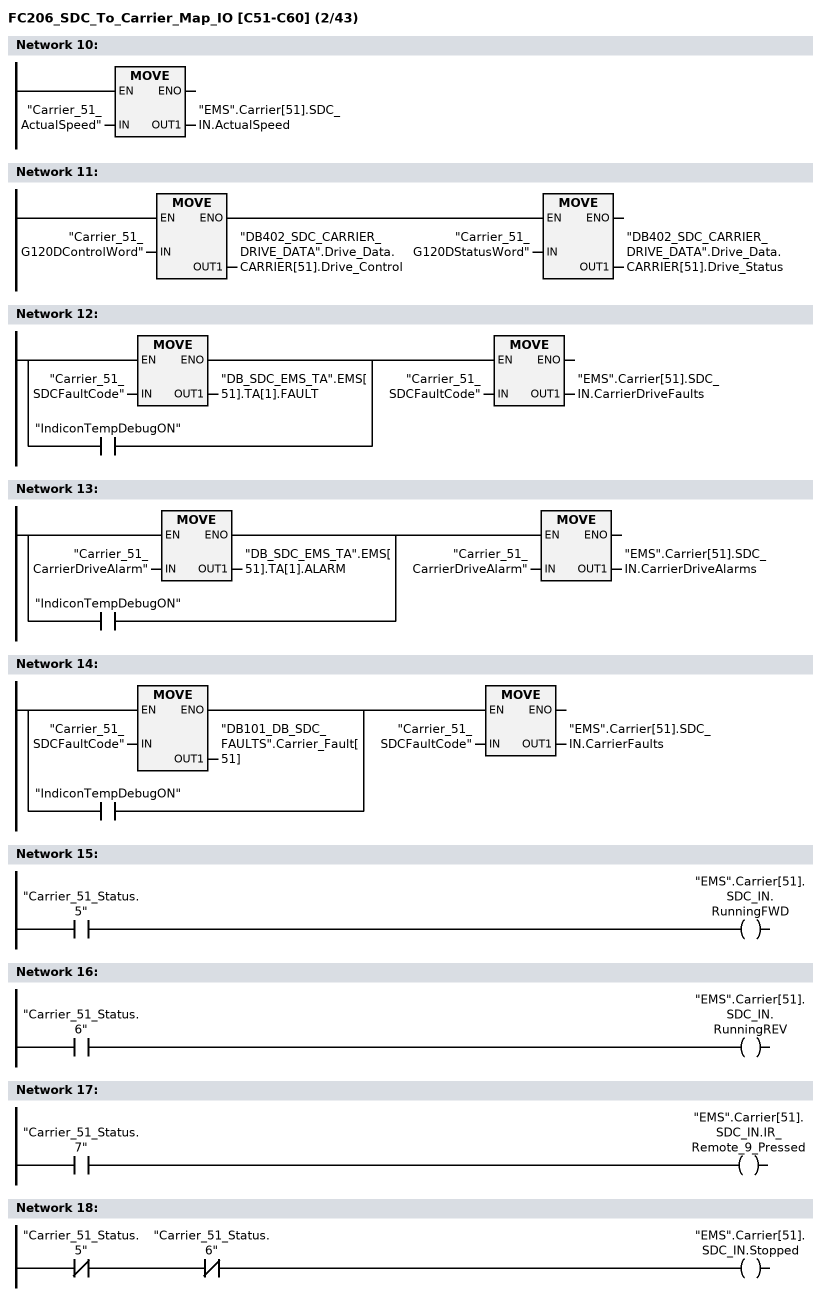
   RUNG wire#powerrail
      Move(in := "Carrier_51_ActualSpeed", out1 => "EMS".Carrier[51].SDC_IN.ActualSpeed)
   END_RUNG
   // the same network as SCL:
   "EMS".Carrier[51].SDC_IN.ActualSpeed := "Carrier_51_ActualSpeed";
END_REGION

REGION Network 11
   RUNG wire#powerrail
      Move(in := "Carrier_51_G120DControlWord", out1 => "DB402_SDC_CARRIER_DRIVE_DATA".Drive_Data.CARRIER[51].Drive_Control)
      Move(in := "Carrier_51_G120DStatusWord", out1 => "DB402_SDC_CARRIER_DRIVE_DATA".Drive_Data.CARRIER[51].Drive_Status)
   END_RUNG
   // the same network as SCL:
   "DB402_SDC_CARRIER_DRIVE_DATA".Drive_Data.CARRIER[51].Drive_Control := "Carrier_51_G120DControlWord";
   "DB402_SDC_CARRIER_DRIVE_DATA".Drive_Data.CARRIER[51].Drive_Status := "Carrier_51_G120DStatusWord";
END_REGION

REGION Network 12
   RUNG wire#powerrail
      Move(in := "Carrier_51_SDCFaultCode", out1 => "DB_SDC_EMS_TA".EMS[51].TA[1].FAULT)
      wire#w1
      Move(in := "Carrier_51_SDCFaultCode", out1 => "EMS".Carrier[51].SDC_IN.CarrierDriveFaults)
   END_RUNG
   RUNG wire#powerrail
      Contact( "IndiconTempDebugON" )
   END_RUNG wire#w1
   // the same network as SCL:
   "DB_SDC_EMS_TA".EMS[51].TA[1].FAULT := "Carrier_51_SDCFaultCode";
   IF TRUE OR "IndiconTempDebugON" THEN
       "EMS".Carrier[51].SDC_IN.CarrierDriveFaults := "Carrier_51_SDCFaultCode";
   END_IF;
END_REGION

REGION Network 13
   RUNG wire#powerrail
      Move(in := "Carrier_51_CarrierDriveAlarm", out1 => "DB_SDC_EMS_TA".EMS[51].TA[1].ALARM)
      wire#w1
      Move(in := "Carrier_51_CarrierDriveAlarm", out1 => "EMS".Carrier[51].SDC_IN.CarrierDriveAlarms)
   END_RUNG
   RUNG wire#powerrail
      Contact( "IndiconTempDebugON" )
   END_RUNG wire#w1
   // the same network as SCL:
   "DB_SDC_EMS_TA".EMS[51].TA[1].ALARM := "Carrier_51_CarrierDriveAlarm";
   IF TRUE OR "IndiconTempDebugON" THEN
       "EMS".Carrier[51].SDC_IN.CarrierDriveAlarms := "Carrier_51_CarrierDriveAlarm";
   END_IF;
END_REGION

REGION Network 14
   RUNG wire#powerrail
      Move(in := "Carrier_51_SDCFaultCode", out1 => "DB101_DB_SDC_FAULTS".Carrier_Fault[51])
      wire#w1
      Move(in := "Carrier_51_SDCFaultCode", out1 => "EMS".Carrier[51].SDC_IN.CarrierFaults)
   END_RUNG
   RUNG wire#powerrail
      Contact( "IndiconTempDebugON" )
   END_RUNG wire#w1
   // the same network as SCL:
   "DB101_DB_SDC_FAULTS".Carrier_Fault[51] := "Carrier_51_SDCFaultCode";
   IF TRUE OR "IndiconTempDebugON" THEN
       "EMS".Carrier[51].SDC_IN.CarrierFaults := "Carrier_51_SDCFaultCode";
   END_IF;
END_REGION

REGION Network 15
   RUNG wire#powerrail
      Contact( "Carrier_51_Status.5" )
      Coil( "EMS".Carrier[51].SDC_IN.RunningFWD )
   END_RUNG
   // the same network as SCL:
   "EMS".Carrier[51].SDC_IN.RunningFWD := "Carrier_51_Status.5";
END_REGION

REGION Network 16
   RUNG wire#powerrail
      Contact( "Carrier_51_Status.6" )
      Coil( "EMS".Carrier[51].SDC_IN.RunningREV )
   END_RUNG
   // the same network as SCL:
   "EMS".Carrier[51].SDC_IN.RunningREV := "Carrier_51_Status.6";
END_REGION

REGION Network 17
   RUNG wire#powerrail
      Contact( "Carrier_51_Status.7" )
      Coil( "EMS".Carrier[51].SDC_IN.IR_Remote_9_Pressed )
   END_RUNG
   // the same network as SCL:
   "EMS".Carrier[51].SDC_IN.IR_Remote_9_Pressed := "Carrier_51_Status.7";
END_REGION

REGION Network 18
   RUNG wire#powerrail
      I_Contact( "Carrier_51_Status.5" )
      I_Contact( "Carrier_51_Status.6" )
      Coil( "EMS".Carrier[51].SDC_IN.Stopped )
   END_RUNG
   // the same network as SCL:
   "EMS".Carrier[51].SDC_IN.Stopped := NOT "Carrier_51_Status.5" AND NOT "Carrier_51_Status.6";
END_REGION

REGION Network 19
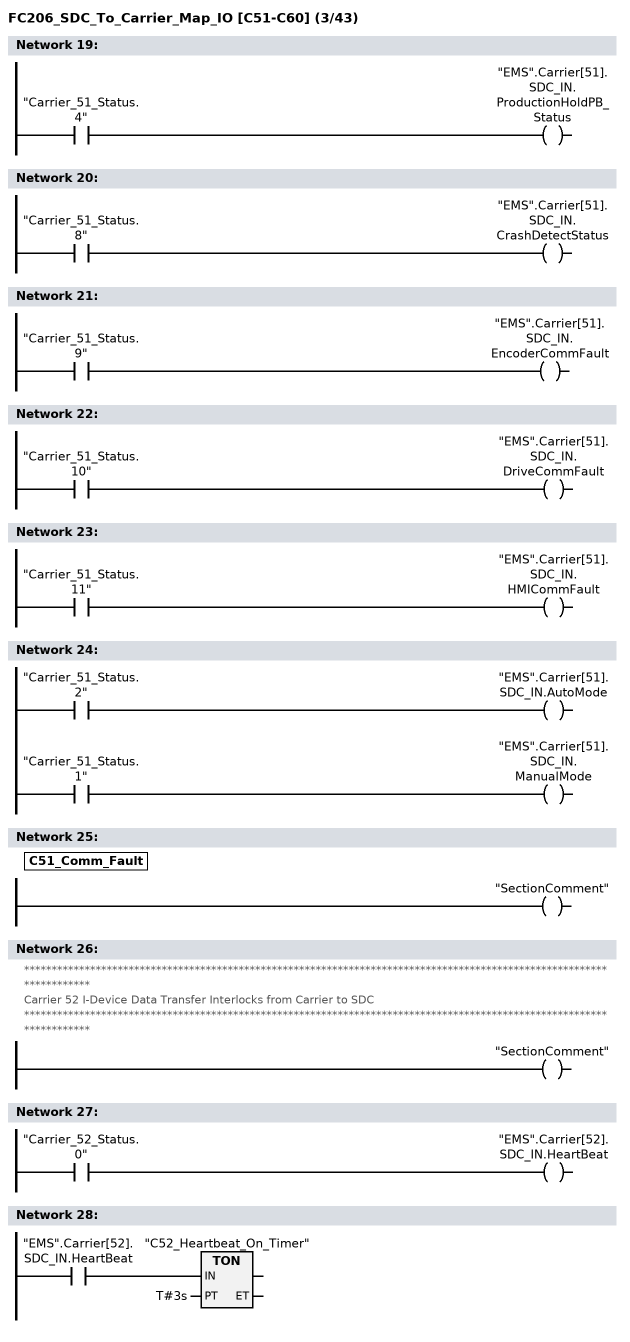
   RUNG wire#powerrail
      Contact( "Carrier_51_Status.4" )
      Coil( "EMS".Carrier[51].SDC_IN.ProductionHoldPB_Status )
   END_RUNG
   // the same network as SCL:
   "EMS".Carrier[51].SDC_IN.ProductionHoldPB_Status := "Carrier_51_Status.4";
END_REGION

REGION Network 20
   RUNG wire#powerrail
      Contact( "Carrier_51_Status.8" )
      Coil( "EMS".Carrier[51].SDC_IN.CrashDetectStatus )
   END_RUNG
   // the same network as SCL:
   "EMS".Carrier[51].SDC_IN.CrashDetectStatus := "Carrier_51_Status.8";
END_REGION

REGION Network 21
   RUNG wire#powerrail
      Contact( "Carrier_51_Status.9" )
      Coil( "EMS".Carrier[51].SDC_IN.EncoderCommFault )
   END_RUNG
   // the same network as SCL:
   "EMS".Carrier[51].SDC_IN.EncoderCommFault := "Carrier_51_Status.9";
END_REGION

REGION Network 22
   RUNG wire#powerrail
      Contact( "Carrier_51_Status.10" )
      Coil( "EMS".Carrier[51].SDC_IN.DriveCommFault )
   END_RUNG
   // the same network as SCL:
   "EMS".Carrier[51].SDC_IN.DriveCommFault := "Carrier_51_Status.10";
END_REGION

REGION Network 23
   RUNG wire#powerrail
      Contact( "Carrier_51_Status.11" )
      Coil( "EMS".Carrier[51].SDC_IN.HMICommFault )
   END_RUNG
   // the same network as SCL:
   "EMS".Carrier[51].SDC_IN.HMICommFault := "Carrier_51_Status.11";
END_REGION

REGION Network 24
   RUNG wire#powerrail
      Contact( "Carrier_51_Status.2" )
      Coil( "EMS".Carrier[51].SDC_IN.AutoMode )
   END_RUNG
   RUNG wire#powerrail
      Contact( "Carrier_51_Status.1" )
      Coil( "EMS".Carrier[51].SDC_IN.ManualMode )
   END_RUNG
   // the same network as SCL:
   "EMS".Carrier[51].SDC_IN.AutoMode := "Carrier_51_Status.2";
   "EMS".Carrier[51].SDC_IN.ManualMode := "Carrier_51_Status.1";
END_REGION

REGION Network 25
   Label( C51_Comm_Fault )
   RUNG wire#powerrail
      Coil( "SectionComment" )
   END_RUNG
   // the same network as SCL:
   C51_Comm_Fault:
   "SectionComment" := TRUE;
END_REGION

REGION Network 26
   // **********************************************************************************************************************
   // 
   // Carrier 52 I-Device Data Transfer Interlocks from Carrier to SDC
   // 
   // **********************************************************************************************************************
   RUNG wire#powerrail
      Coil( "SectionComment" )
   END_RUNG
   // the same network as SCL:
   "SectionComment" := TRUE;
END_REGION

REGION Network 27
   RUNG wire#powerrail
      Contact( "Carrier_52_Status.0" )
      Coil( "EMS".Carrier[52].SDC_IN.HeartBeat )
   END_RUNG
   // the same network as SCL:
   "EMS".Carrier[52].SDC_IN.HeartBeat := "Carrier_52_Status.0";
END_REGION

REGION Network 28
   "C52_Heartbeat_On_Timer".TON(IN := "EMS".Carrier[52].SDC_IN.HeartBeat, PT := T#3s);
END_REGION

REGION Network 29
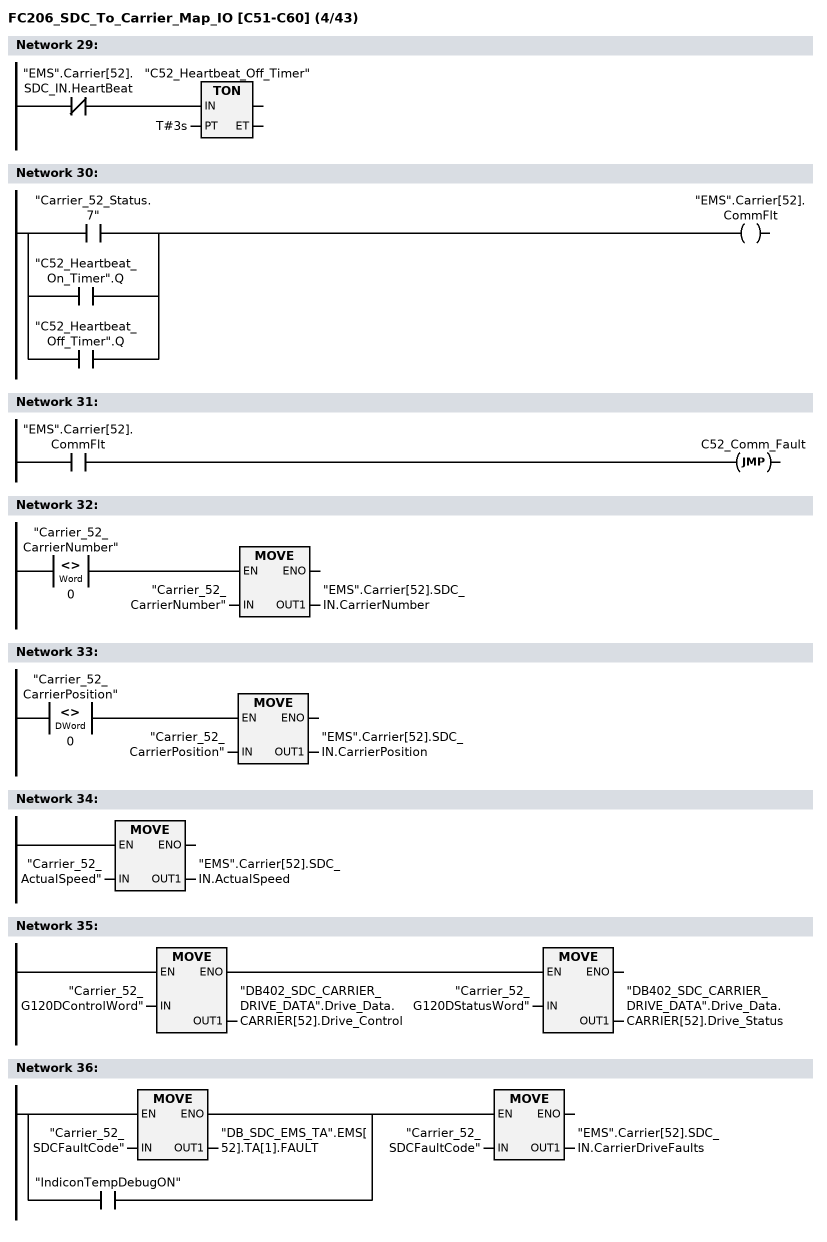
   "C52_Heartbeat_Off_Timer".TON(IN := NOT "EMS".Carrier[52].SDC_IN.HeartBeat, PT := T#3s);
END_REGION

REGION Network 30
   RUNG wire#powerrail
      Contact( "Carrier_52_Status.7" )
      wire#w1
      Coil( "EMS".Carrier[52].CommFlt )
   END_RUNG
   RUNG wire#powerrail
      Contact( "C52_Heartbeat_On_Timer".Q )
   END_RUNG wire#w1
   RUNG wire#powerrail
      Contact( "C52_Heartbeat_Off_Timer".Q )
   END_RUNG wire#w1
   // the same network as SCL:
   "EMS".Carrier[52].CommFlt := "Carrier_52_Status.7" OR "C52_Heartbeat_On_Timer".Q OR "C52_Heartbeat_Off_Timer".Q;
END_REGION

REGION Network 31
   RUNG wire#powerrail
      Contact( "EMS".Carrier[52].CommFlt )
      JumpCoil( C52_Comm_Fault )
   END_RUNG
   // the same network as SCL:
   IF "EMS".Carrier[52].CommFlt THEN GOTO C52_Comm_Fault; END_IF;
END_REGION

REGION Network 32
   RUNG wire#powerrail
      { S7_Templates := "SrcType := Word" } NE_Contact(in1 := "Carrier_52_CarrierNumber", in2 := 0)
      Move(in := "Carrier_52_CarrierNumber", out1 => "EMS".Carrier[52].SDC_IN.CarrierNumber)
   END_RUNG
   // the same network as SCL:
   IF "Carrier_52_CarrierNumber" <> 0 THEN
       "EMS".Carrier[52].SDC_IN.CarrierNumber := "Carrier_52_CarrierNumber";
   END_IF;
END_REGION

REGION Network 33
   RUNG wire#powerrail
      { S7_Templates := "SrcType := DWord" } NE_Contact(in1 := "Carrier_52_CarrierPosition", in2 := 0)
      Move(in := "Carrier_52_CarrierPosition", out1 => "EMS".Carrier[52].SDC_IN.CarrierPosition)
   END_RUNG
   // the same network as SCL:
   IF "Carrier_52_CarrierPosition" <> 0 THEN
       "EMS".Carrier[52].SDC_IN.CarrierPosition := "Carrier_52_CarrierPosition";
   END_IF;
END_REGION

REGION Network 34
   RUNG wire#powerrail
      Move(in := "Carrier_52_ActualSpeed", out1 => "EMS".Carrier[52].SDC_IN.ActualSpeed)
   END_RUNG
   // the same network as SCL:
   "EMS".Carrier[52].SDC_IN.ActualSpeed := "Carrier_52_ActualSpeed";
END_REGION

REGION Network 35
   RUNG wire#powerrail
      Move(in := "Carrier_52_G120DControlWord", out1 => "DB402_SDC_CARRIER_DRIVE_DATA".Drive_Data.CARRIER[52].Drive_Control)
      Move(in := "Carrier_52_G120DStatusWord", out1 => "DB402_SDC_CARRIER_DRIVE_DATA".Drive_Data.CARRIER[52].Drive_Status)
   END_RUNG
   // the same network as SCL:
   "DB402_SDC_CARRIER_DRIVE_DATA".Drive_Data.CARRIER[52].Drive_Control := "Carrier_52_G120DControlWord";
   "DB402_SDC_CARRIER_DRIVE_DATA".Drive_Data.CARRIER[52].Drive_Status := "Carrier_52_G120DStatusWord";
END_REGION

REGION Network 36
   RUNG wire#powerrail
      Move(in := "Carrier_52_SDCFaultCode", out1 => "DB_SDC_EMS_TA".EMS[52].TA[1].FAULT)
      wire#w1
      Move(in := "Carrier_52_SDCFaultCode", out1 => "EMS".Carrier[52].SDC_IN.CarrierDriveFaults)
   END_RUNG
   RUNG wire#powerrail
      Contact( "IndiconTempDebugON" )
   END_RUNG wire#w1
   // the same network as SCL:
   "DB_SDC_EMS_TA".EMS[52].TA[1].FAULT := "Carrier_52_SDCFaultCode";
   IF TRUE OR "IndiconTempDebugON" THEN
       "EMS".Carrier[52].SDC_IN.CarrierDriveFaults := "Carrier_52_SDCFaultCode";
   END_IF;
END_REGION

REGION Network 37
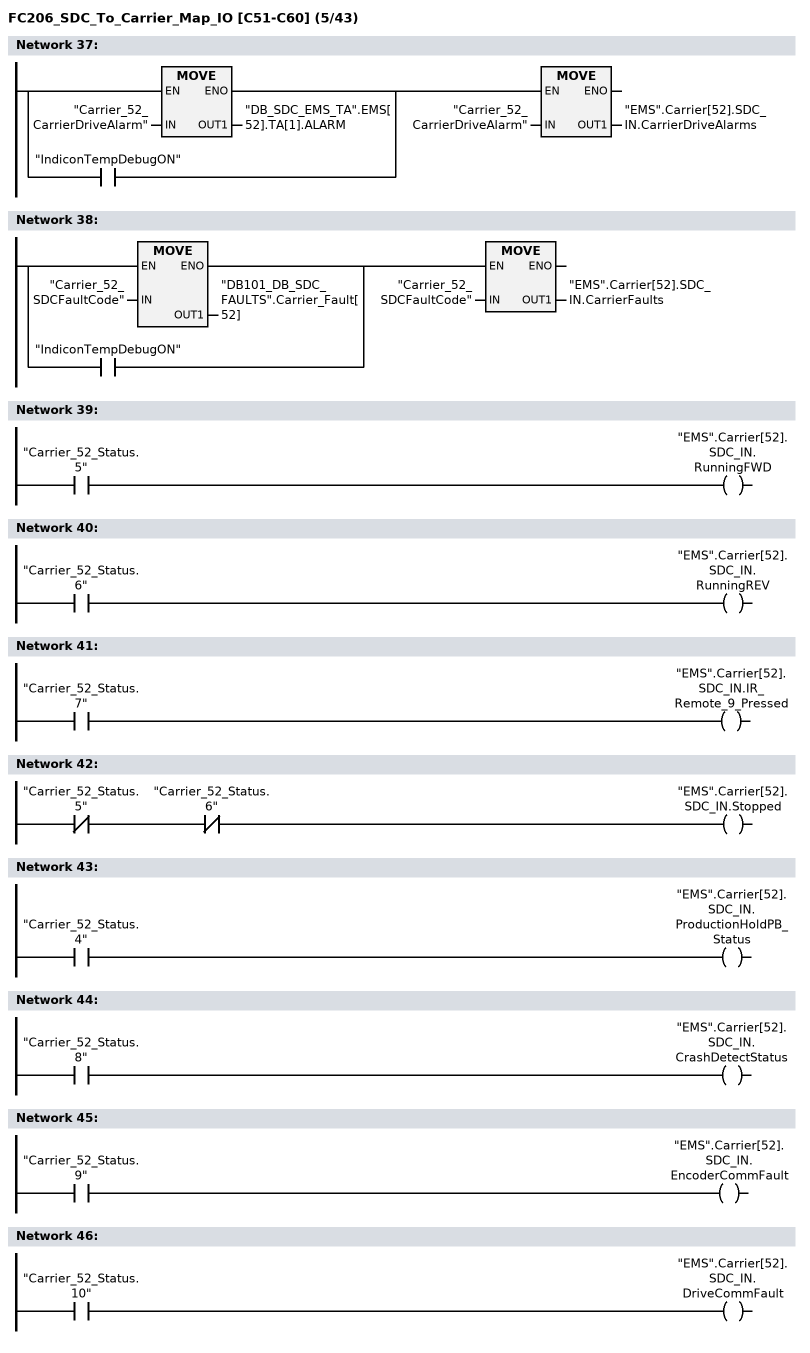
   RUNG wire#powerrail
      Move(in := "Carrier_52_CarrierDriveAlarm", out1 => "DB_SDC_EMS_TA".EMS[52].TA[1].ALARM)
      wire#w1
      Move(in := "Carrier_52_CarrierDriveAlarm", out1 => "EMS".Carrier[52].SDC_IN.CarrierDriveAlarms)
   END_RUNG
   RUNG wire#powerrail
      Contact( "IndiconTempDebugON" )
   END_RUNG wire#w1
   // the same network as SCL:
   "DB_SDC_EMS_TA".EMS[52].TA[1].ALARM := "Carrier_52_CarrierDriveAlarm";
   IF TRUE OR "IndiconTempDebugON" THEN
       "EMS".Carrier[52].SDC_IN.CarrierDriveAlarms := "Carrier_52_CarrierDriveAlarm";
   END_IF;
END_REGION

REGION Network 38
   RUNG wire#powerrail
      Move(in := "Carrier_52_SDCFaultCode", out1 => "DB101_DB_SDC_FAULTS".Carrier_Fault[52])
      wire#w1
      Move(in := "Carrier_52_SDCFaultCode", out1 => "EMS".Carrier[52].SDC_IN.CarrierFaults)
   END_RUNG
   RUNG wire#powerrail
      Contact( "IndiconTempDebugON" )
   END_RUNG wire#w1
   // the same network as SCL:
   "DB101_DB_SDC_FAULTS".Carrier_Fault[52] := "Carrier_52_SDCFaultCode";
   IF TRUE OR "IndiconTempDebugON" THEN
       "EMS".Carrier[52].SDC_IN.CarrierFaults := "Carrier_52_SDCFaultCode";
   END_IF;
END_REGION

REGION Network 39
   RUNG wire#powerrail
      Contact( "Carrier_52_Status.5" )
      Coil( "EMS".Carrier[52].SDC_IN.RunningFWD )
   END_RUNG
   // the same network as SCL:
   "EMS".Carrier[52].SDC_IN.RunningFWD := "Carrier_52_Status.5";
END_REGION

REGION Network 40
   RUNG wire#powerrail
      Contact( "Carrier_52_Status.6" )
      Coil( "EMS".Carrier[52].SDC_IN.RunningREV )
   END_RUNG
   // the same network as SCL:
   "EMS".Carrier[52].SDC_IN.RunningREV := "Carrier_52_Status.6";
END_REGION

REGION Network 41
   RUNG wire#powerrail
      Contact( "Carrier_52_Status.7" )
      Coil( "EMS".Carrier[52].SDC_IN.IR_Remote_9_Pressed )
   END_RUNG
   // the same network as SCL:
   "EMS".Carrier[52].SDC_IN.IR_Remote_9_Pressed := "Carrier_52_Status.7";
END_REGION

REGION Network 42
   RUNG wire#powerrail
      I_Contact( "Carrier_52_Status.5" )
      I_Contact( "Carrier_52_Status.6" )
      Coil( "EMS".Carrier[52].SDC_IN.Stopped )
   END_RUNG
   // the same network as SCL:
   "EMS".Carrier[52].SDC_IN.Stopped := NOT "Carrier_52_Status.5" AND NOT "Carrier_52_Status.6";
END_REGION

REGION Network 43
   RUNG wire#powerrail
      Contact( "Carrier_52_Status.4" )
      Coil( "EMS".Carrier[52].SDC_IN.ProductionHoldPB_Status )
   END_RUNG
   // the same network as SCL:
   "EMS".Carrier[52].SDC_IN.ProductionHoldPB_Status := "Carrier_52_Status.4";
END_REGION

REGION Network 44
   RUNG wire#powerrail
      Contact( "Carrier_52_Status.8" )
      Coil( "EMS".Carrier[52].SDC_IN.CrashDetectStatus )
   END_RUNG
   // the same network as SCL:
   "EMS".Carrier[52].SDC_IN.CrashDetectStatus := "Carrier_52_Status.8";
END_REGION

REGION Network 45
   RUNG wire#powerrail
      Contact( "Carrier_52_Status.9" )
      Coil( "EMS".Carrier[52].SDC_IN.EncoderCommFault )
   END_RUNG
   // the same network as SCL:
   "EMS".Carrier[52].SDC_IN.EncoderCommFault := "Carrier_52_Status.9";
END_REGION

REGION Network 46
   RUNG wire#powerrail
      Contact( "Carrier_52_Status.10" )
      Coil( "EMS".Carrier[52].SDC_IN.DriveCommFault )
   END_RUNG
   // the same network as SCL:
   "EMS".Carrier[52].SDC_IN.DriveCommFault := "Carrier_52_Status.10";
END_REGION

REGION Network 47
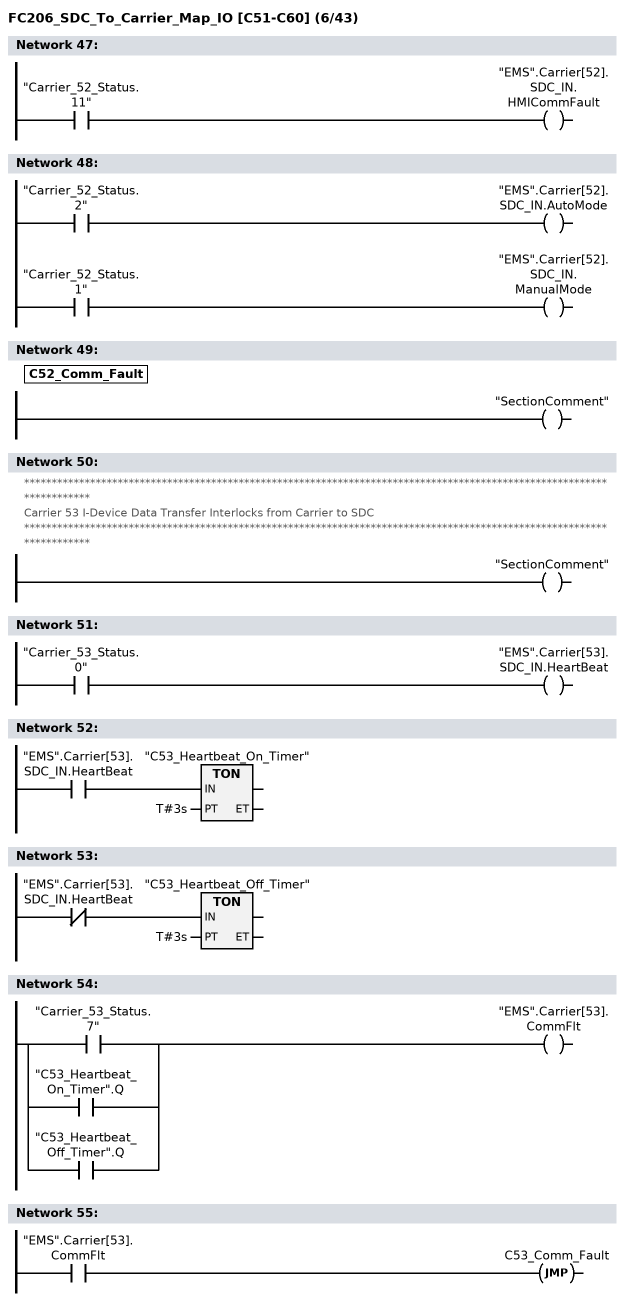
   RUNG wire#powerrail
      Contact( "Carrier_52_Status.11" )
      Coil( "EMS".Carrier[52].SDC_IN.HMICommFault )
   END_RUNG
   // the same network as SCL:
   "EMS".Carrier[52].SDC_IN.HMICommFault := "Carrier_52_Status.11";
END_REGION

REGION Network 48
   RUNG wire#powerrail
      Contact( "Carrier_52_Status.2" )
      Coil( "EMS".Carrier[52].SDC_IN.AutoMode )
   END_RUNG
   RUNG wire#powerrail
      Contact( "Carrier_52_Status.1" )
      Coil( "EMS".Carrier[52].SDC_IN.ManualMode )
   END_RUNG
   // the same network as SCL:
   "EMS".Carrier[52].SDC_IN.AutoMode := "Carrier_52_Status.2";
   "EMS".Carrier[52].SDC_IN.ManualMode := "Carrier_52_Status.1";
END_REGION

REGION Network 49
   Label( C52_Comm_Fault )
   RUNG wire#powerrail
      Coil( "SectionComment" )
   END_RUNG
   // the same network as SCL:
   C52_Comm_Fault:
   "SectionComment" := TRUE;
END_REGION

REGION Network 50
   // **********************************************************************************************************************
   // 
   // Carrier 53 I-Device Data Transfer Interlocks from Carrier to SDC
   // 
   // **********************************************************************************************************************
   RUNG wire#powerrail
      Coil( "SectionComment" )
   END_RUNG
   // the same network as SCL:
   "SectionComment" := TRUE;
END_REGION

REGION Network 51
   RUNG wire#powerrail
      Contact( "Carrier_53_Status.0" )
      Coil( "EMS".Carrier[53].SDC_IN.HeartBeat )
   END_RUNG
   // the same network as SCL:
   "EMS".Carrier[53].SDC_IN.HeartBeat := "Carrier_53_Status.0";
END_REGION

REGION Network 52
   "C53_Heartbeat_On_Timer".TON(IN := "EMS".Carrier[53].SDC_IN.HeartBeat, PT := T#3s);
END_REGION

REGION Network 53
   "C53_Heartbeat_Off_Timer".TON(IN := NOT "EMS".Carrier[53].SDC_IN.HeartBeat, PT := T#3s);
END_REGION

REGION Network 54
   RUNG wire#powerrail
      Contact( "Carrier_53_Status.7" )
      wire#w1
      Coil( "EMS".Carrier[53].CommFlt )
   END_RUNG
   RUNG wire#powerrail
      Contact( "C53_Heartbeat_On_Timer".Q )
   END_RUNG wire#w1
   RUNG wire#powerrail
      Contact( "C53_Heartbeat_Off_Timer".Q )
   END_RUNG wire#w1
   // the same network as SCL:
   "EMS".Carrier[53].CommFlt := "Carrier_53_Status.7" OR "C53_Heartbeat_On_Timer".Q OR "C53_Heartbeat_Off_Timer".Q;
END_REGION

REGION Network 55
   RUNG wire#powerrail
      Contact( "EMS".Carrier[53].CommFlt )
      JumpCoil( C53_Comm_Fault )
   END_RUNG
   // the same network as SCL:
   IF "EMS".Carrier[53].CommFlt THEN GOTO C53_Comm_Fault; END_IF;
END_REGION

REGION Network 56
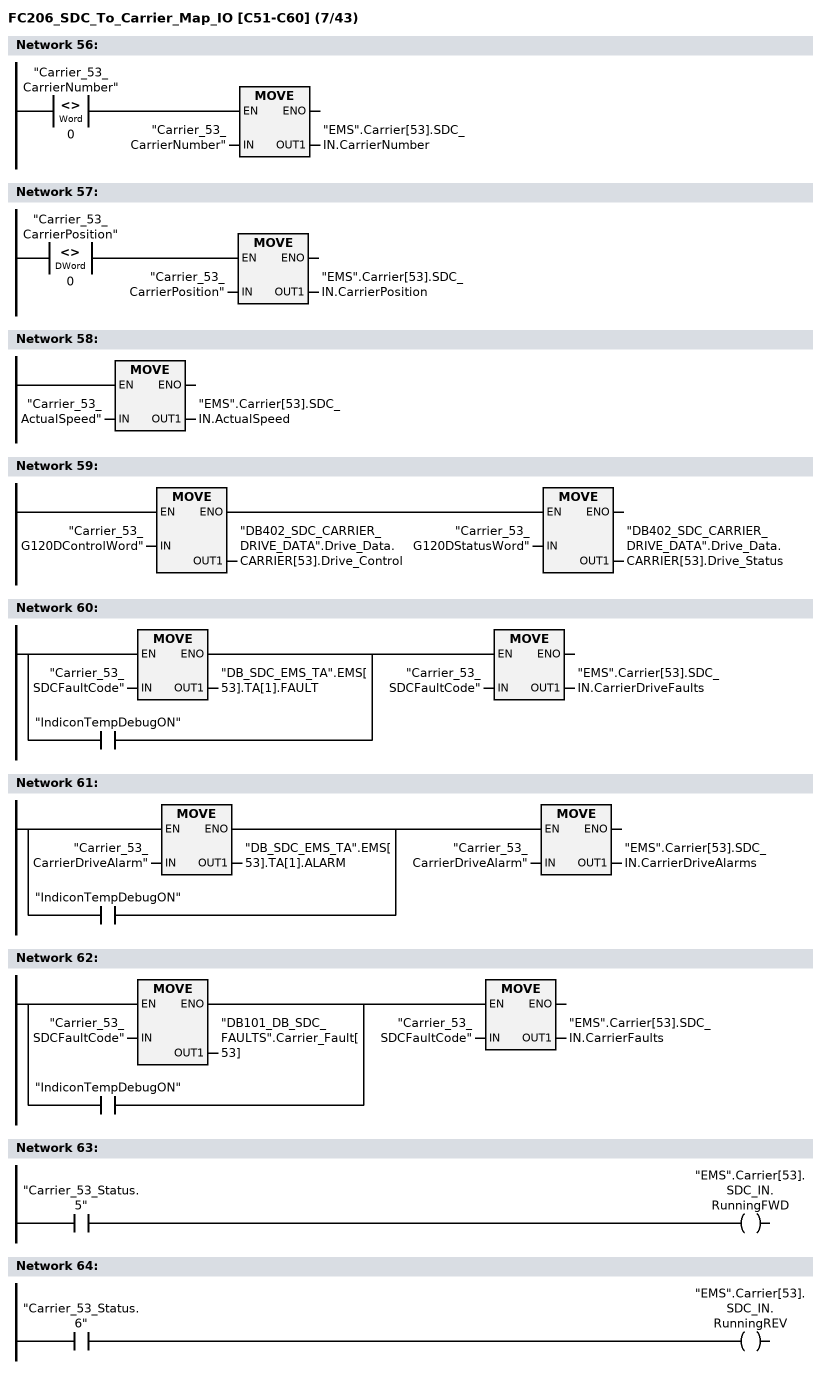
   RUNG wire#powerrail
      { S7_Templates := "SrcType := Word" } NE_Contact(in1 := "Carrier_53_CarrierNumber", in2 := 0)
      Move(in := "Carrier_53_CarrierNumber", out1 => "EMS".Carrier[53].SDC_IN.CarrierNumber)
   END_RUNG
   // the same network as SCL:
   IF "Carrier_53_CarrierNumber" <> 0 THEN
       "EMS".Carrier[53].SDC_IN.CarrierNumber := "Carrier_53_CarrierNumber";
   END_IF;
END_REGION

REGION Network 57
   RUNG wire#powerrail
      { S7_Templates := "SrcType := DWord" } NE_Contact(in1 := "Carrier_53_CarrierPosition", in2 := 0)
      Move(in := "Carrier_53_CarrierPosition", out1 => "EMS".Carrier[53].SDC_IN.CarrierPosition)
   END_RUNG
   // the same network as SCL:
   IF "Carrier_53_CarrierPosition" <> 0 THEN
       "EMS".Carrier[53].SDC_IN.CarrierPosition := "Carrier_53_CarrierPosition";
   END_IF;
END_REGION

REGION Network 58
   RUNG wire#powerrail
      Move(in := "Carrier_53_ActualSpeed", out1 => "EMS".Carrier[53].SDC_IN.ActualSpeed)
   END_RUNG
   // the same network as SCL:
   "EMS".Carrier[53].SDC_IN.ActualSpeed := "Carrier_53_ActualSpeed";
END_REGION

REGION Network 59
   RUNG wire#powerrail
      Move(in := "Carrier_53_G120DControlWord", out1 => "DB402_SDC_CARRIER_DRIVE_DATA".Drive_Data.CARRIER[53].Drive_Control)
      Move(in := "Carrier_53_G120DStatusWord", out1 => "DB402_SDC_CARRIER_DRIVE_DATA".Drive_Data.CARRIER[53].Drive_Status)
   END_RUNG
   // the same network as SCL:
   "DB402_SDC_CARRIER_DRIVE_DATA".Drive_Data.CARRIER[53].Drive_Control := "Carrier_53_G120DControlWord";
   "DB402_SDC_CARRIER_DRIVE_DATA".Drive_Data.CARRIER[53].Drive_Status := "Carrier_53_G120DStatusWord";
END_REGION

REGION Network 60
   RUNG wire#powerrail
      Move(in := "Carrier_53_SDCFaultCode", out1 => "DB_SDC_EMS_TA".EMS[53].TA[1].FAULT)
      wire#w1
      Move(in := "Carrier_53_SDCFaultCode", out1 => "EMS".Carrier[53].SDC_IN.CarrierDriveFaults)
   END_RUNG
   RUNG wire#powerrail
      Contact( "IndiconTempDebugON" )
   END_RUNG wire#w1
   // the same network as SCL:
   "DB_SDC_EMS_TA".EMS[53].TA[1].FAULT := "Carrier_53_SDCFaultCode";
   IF TRUE OR "IndiconTempDebugON" THEN
       "EMS".Carrier[53].SDC_IN.CarrierDriveFaults := "Carrier_53_SDCFaultCode";
   END_IF;
END_REGION

REGION Network 61
   RUNG wire#powerrail
      Move(in := "Carrier_53_CarrierDriveAlarm", out1 => "DB_SDC_EMS_TA".EMS[53].TA[1].ALARM)
      wire#w1
      Move(in := "Carrier_53_CarrierDriveAlarm", out1 => "EMS".Carrier[53].SDC_IN.CarrierDriveAlarms)
   END_RUNG
   RUNG wire#powerrail
      Contact( "IndiconTempDebugON" )
   END_RUNG wire#w1
   // the same network as SCL:
   "DB_SDC_EMS_TA".EMS[53].TA[1].ALARM := "Carrier_53_CarrierDriveAlarm";
   IF TRUE OR "IndiconTempDebugON" THEN
       "EMS".Carrier[53].SDC_IN.CarrierDriveAlarms := "Carrier_53_CarrierDriveAlarm";
   END_IF;
END_REGION

REGION Network 62
   RUNG wire#powerrail
      Move(in := "Carrier_53_SDCFaultCode", out1 => "DB101_DB_SDC_FAULTS".Carrier_Fault[53])
      wire#w1
      Move(in := "Carrier_53_SDCFaultCode", out1 => "EMS".Carrier[53].SDC_IN.CarrierFaults)
   END_RUNG
   RUNG wire#powerrail
      Contact( "IndiconTempDebugON" )
   END_RUNG wire#w1
   // the same network as SCL:
   "DB101_DB_SDC_FAULTS".Carrier_Fault[53] := "Carrier_53_SDCFaultCode";
   IF TRUE OR "IndiconTempDebugON" THEN
       "EMS".Carrier[53].SDC_IN.CarrierFaults := "Carrier_53_SDCFaultCode";
   END_IF;
END_REGION

REGION Network 63
   RUNG wire#powerrail
      Contact( "Carrier_53_Status.5" )
      Coil( "EMS".Carrier[53].SDC_IN.RunningFWD )
   END_RUNG
   // the same network as SCL:
   "EMS".Carrier[53].SDC_IN.RunningFWD := "Carrier_53_Status.5";
END_REGION

REGION Network 64
   RUNG wire#powerrail
      Contact( "Carrier_53_Status.6" )
      Coil( "EMS".Carrier[53].SDC_IN.RunningREV )
   END_RUNG
   // the same network as SCL:
   "EMS".Carrier[53].SDC_IN.RunningREV := "Carrier_53_Status.6";
END_REGION

REGION Network 65
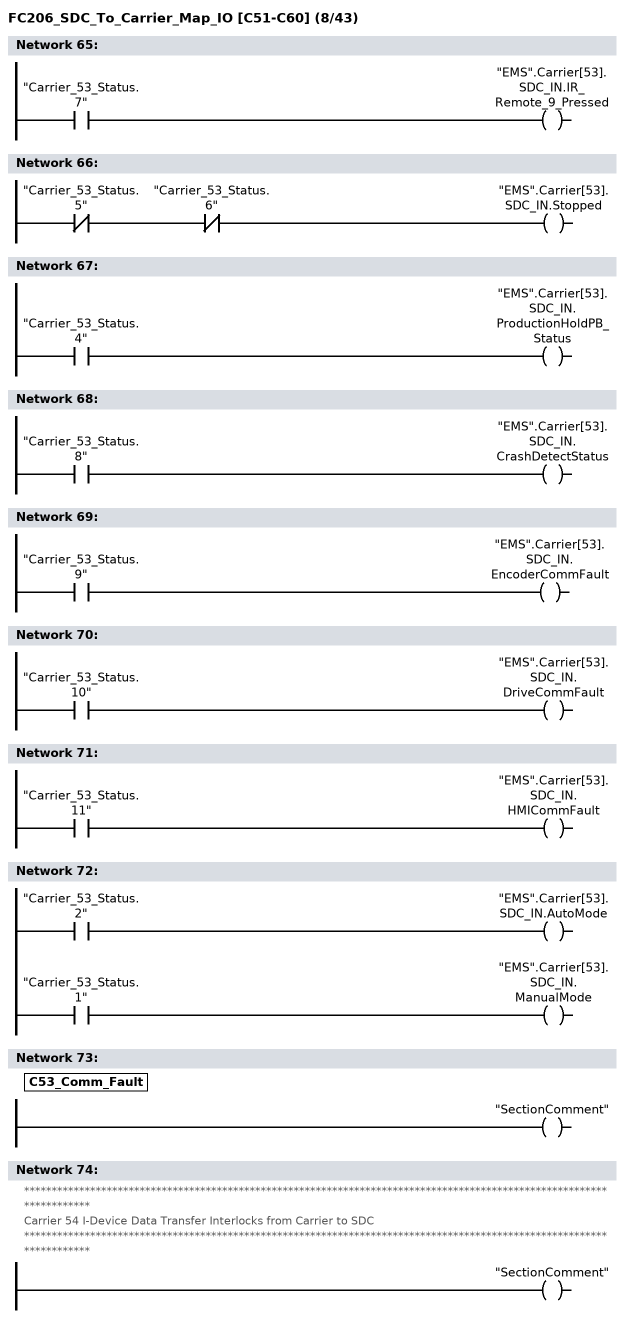
   RUNG wire#powerrail
      Contact( "Carrier_53_Status.7" )
      Coil( "EMS".Carrier[53].SDC_IN.IR_Remote_9_Pressed )
   END_RUNG
   // the same network as SCL:
   "EMS".Carrier[53].SDC_IN.IR_Remote_9_Pressed := "Carrier_53_Status.7";
END_REGION

REGION Network 66
   RUNG wire#powerrail
      I_Contact( "Carrier_53_Status.5" )
      I_Contact( "Carrier_53_Status.6" )
      Coil( "EMS".Carrier[53].SDC_IN.Stopped )
   END_RUNG
   // the same network as SCL:
   "EMS".Carrier[53].SDC_IN.Stopped := NOT "Carrier_53_Status.5" AND NOT "Carrier_53_Status.6";
END_REGION

REGION Network 67
   RUNG wire#powerrail
      Contact( "Carrier_53_Status.4" )
      Coil( "EMS".Carrier[53].SDC_IN.ProductionHoldPB_Status )
   END_RUNG
   // the same network as SCL:
   "EMS".Carrier[53].SDC_IN.ProductionHoldPB_Status := "Carrier_53_Status.4";
END_REGION

REGION Network 68
   RUNG wire#powerrail
      Contact( "Carrier_53_Status.8" )
      Coil( "EMS".Carrier[53].SDC_IN.CrashDetectStatus )
   END_RUNG
   // the same network as SCL:
   "EMS".Carrier[53].SDC_IN.CrashDetectStatus := "Carrier_53_Status.8";
END_REGION

REGION Network 69
   RUNG wire#powerrail
      Contact( "Carrier_53_Status.9" )
      Coil( "EMS".Carrier[53].SDC_IN.EncoderCommFault )
   END_RUNG
   // the same network as SCL:
   "EMS".Carrier[53].SDC_IN.EncoderCommFault := "Carrier_53_Status.9";
END_REGION

REGION Network 70
   RUNG wire#powerrail
      Contact( "Carrier_53_Status.10" )
      Coil( "EMS".Carrier[53].SDC_IN.DriveCommFault )
   END_RUNG
   // the same network as SCL:
   "EMS".Carrier[53].SDC_IN.DriveCommFault := "Carrier_53_Status.10";
END_REGION

REGION Network 71
   RUNG wire#powerrail
      Contact( "Carrier_53_Status.11" )
      Coil( "EMS".Carrier[53].SDC_IN.HMICommFault )
   END_RUNG
   // the same network as SCL:
   "EMS".Carrier[53].SDC_IN.HMICommFault := "Carrier_53_Status.11";
END_REGION

REGION Network 72
   RUNG wire#powerrail
      Contact( "Carrier_53_Status.2" )
      Coil( "EMS".Carrier[53].SDC_IN.AutoMode )
   END_RUNG
   RUNG wire#powerrail
      Contact( "Carrier_53_Status.1" )
      Coil( "EMS".Carrier[53].SDC_IN.ManualMode )
   END_RUNG
   // the same network as SCL:
   "EMS".Carrier[53].SDC_IN.AutoMode := "Carrier_53_Status.2";
   "EMS".Carrier[53].SDC_IN.ManualMode := "Carrier_53_Status.1";
END_REGION

REGION Network 73
   Label( C53_Comm_Fault )
   RUNG wire#powerrail
      Coil( "SectionComment" )
   END_RUNG
   // the same network as SCL:
   C53_Comm_Fault:
   "SectionComment" := TRUE;
END_REGION

REGION Network 74
   // **********************************************************************************************************************
   // 
   // Carrier 54 I-Device Data Transfer Interlocks from Carrier to SDC
   // 
   // **********************************************************************************************************************
   RUNG wire#powerrail
      Coil( "SectionComment" )
   END_RUNG
   // the same network as SCL:
   "SectionComment" := TRUE;
END_REGION

REGION Network 75
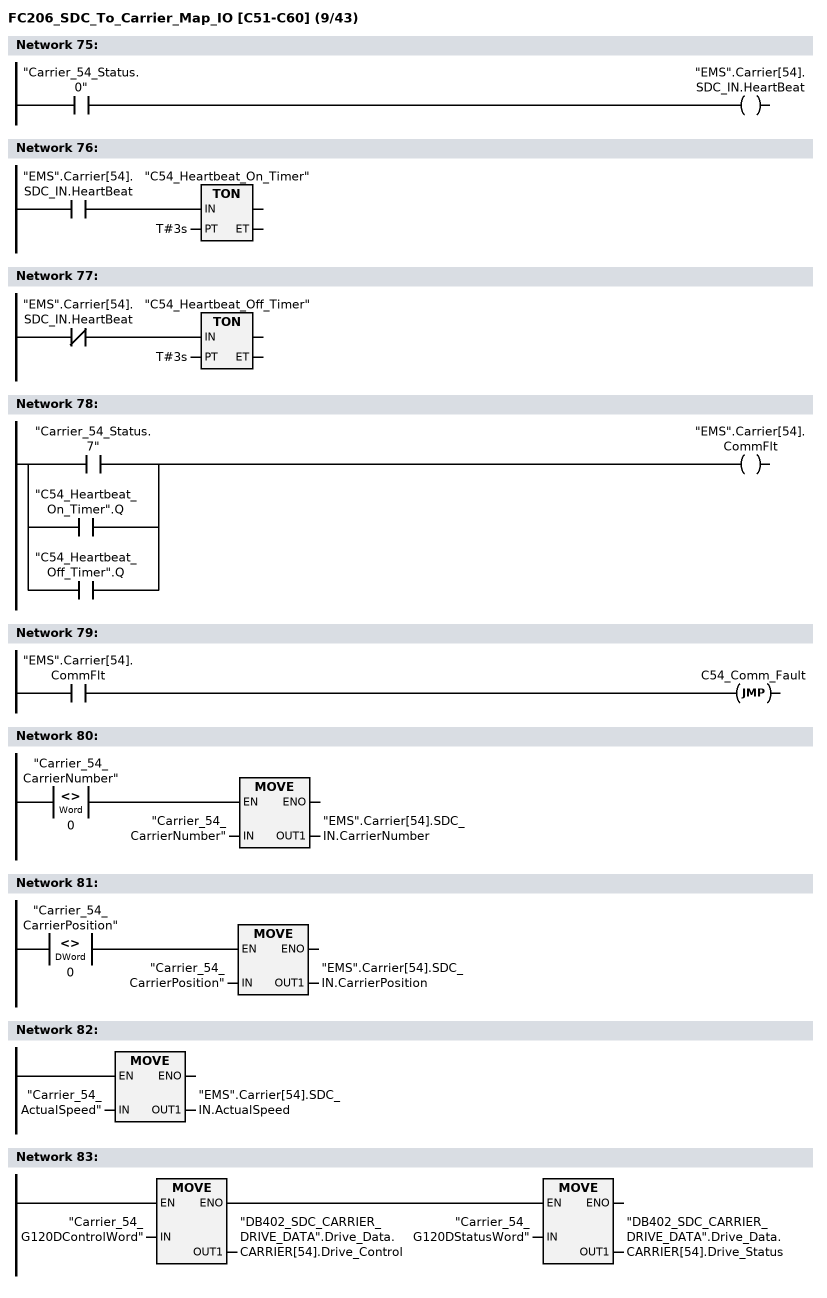
   RUNG wire#powerrail
      Contact( "Carrier_54_Status.0" )
      Coil( "EMS".Carrier[54].SDC_IN.HeartBeat )
   END_RUNG
   // the same network as SCL:
   "EMS".Carrier[54].SDC_IN.HeartBeat := "Carrier_54_Status.0";
END_REGION

REGION Network 76
   "C54_Heartbeat_On_Timer".TON(IN := "EMS".Carrier[54].SDC_IN.HeartBeat, PT := T#3s);
END_REGION

REGION Network 77
   "C54_Heartbeat_Off_Timer".TON(IN := NOT "EMS".Carrier[54].SDC_IN.HeartBeat, PT := T#3s);
END_REGION

REGION Network 78
   RUNG wire#powerrail
      Contact( "Carrier_54_Status.7" )
      wire#w1
      Coil( "EMS".Carrier[54].CommFlt )
   END_RUNG
   RUNG wire#powerrail
      Contact( "C54_Heartbeat_On_Timer".Q )
   END_RUNG wire#w1
   RUNG wire#powerrail
      Contact( "C54_Heartbeat_Off_Timer".Q )
   END_RUNG wire#w1
   // the same network as SCL:
   "EMS".Carrier[54].CommFlt := "Carrier_54_Status.7" OR "C54_Heartbeat_On_Timer".Q OR "C54_Heartbeat_Off_Timer".Q;
END_REGION

REGION Network 79
   RUNG wire#powerrail
      Contact( "EMS".Carrier[54].CommFlt )
      JumpCoil( C54_Comm_Fault )
   END_RUNG
   // the same network as SCL:
   IF "EMS".Carrier[54].CommFlt THEN GOTO C54_Comm_Fault; END_IF;
END_REGION

REGION Network 80
   RUNG wire#powerrail
      { S7_Templates := "SrcType := Word" } NE_Contact(in1 := "Carrier_54_CarrierNumber", in2 := 0)
      Move(in := "Carrier_54_CarrierNumber", out1 => "EMS".Carrier[54].SDC_IN.CarrierNumber)
   END_RUNG
   // the same network as SCL:
   IF "Carrier_54_CarrierNumber" <> 0 THEN
       "EMS".Carrier[54].SDC_IN.CarrierNumber := "Carrier_54_CarrierNumber";
   END_IF;
END_REGION

REGION Network 81
   RUNG wire#powerrail
      { S7_Templates := "SrcType := DWord" } NE_Contact(in1 := "Carrier_54_CarrierPosition", in2 := 0)
      Move(in := "Carrier_54_CarrierPosition", out1 => "EMS".Carrier[54].SDC_IN.CarrierPosition)
   END_RUNG
   // the same network as SCL:
   IF "Carrier_54_CarrierPosition" <> 0 THEN
       "EMS".Carrier[54].SDC_IN.CarrierPosition := "Carrier_54_CarrierPosition";
   END_IF;
END_REGION

REGION Network 82
   RUNG wire#powerrail
      Move(in := "Carrier_54_ActualSpeed", out1 => "EMS".Carrier[54].SDC_IN.ActualSpeed)
   END_RUNG
   // the same network as SCL:
   "EMS".Carrier[54].SDC_IN.ActualSpeed := "Carrier_54_ActualSpeed";
END_REGION
